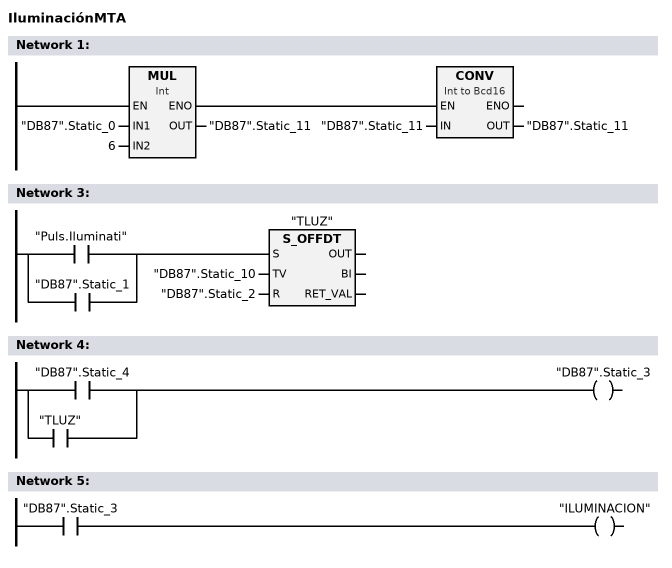
   RUNG wire#powerrail
      { S7_Templates := "SrcType := Int"; S7_GenerateENO := "TRUE" } Mul(in1 := "DB87".Static_0, in2 := 6, out => "DB87".Static_11)
      { S7_Templates := "[SrcType := Int, DestType := Bcd16]"; S7_GenerateENO := "TRUE" } Convert(in := "DB87".Static_11, out => "DB87".Static_11)
   END_RUNG
   // the same network as SCL:
   // ENO of a box is taken as its EN; it also drops when the box reports an error
   "DB87".Static_11 := "DB87".Static_0 * 6;
   "DB87".Static_11 := INT_TO_BCD16("DB87".Static_11);
END_REGION

REGION Network 2 (STL)
         L     12288;
         L     "DB87".Static_11;
         OW;
         T     "DB87".Static_10;
         NOP   0;
END_REGION

REGION Network 3
   RUNG wire#powerrail
      Contact( "Puls.Iluminati" )
      wire#w1
      S_OFFDT(T_NO := "TLUZ", TV := "DB87".Static_10, R := "DB87".Static_2, BI =>, RET_VAL =>)
   END_RUNG
   RUNG wire#powerrail
      Contact( "DB87".Static_1 )
   END_RUNG wire#w1
   // the same network as SCL:
   #_s5time1 := S_OFFDT(T_NO := "TLUZ",
                        S := "Puls.Iluminati" OR "DB87".Static_1,
                        TV := "DB87".Static_10,
                        R := "DB87".Static_2);
END_REGION

REGION Network 4
   RUNG wire#powerrail
      Contact( "DB87".Static_4 )
      wire#w1
      Coil( "DB87".Static_3 )
   END_RUNG
   RUNG wire#powerrail
      Contact( "TLUZ" )
   END_RUNG wire#w1
   // the same network as SCL:
   "DB87".Static_3 := "DB87".Static_4 OR "TLUZ";
END_REGION

REGION Network 5
   RUNG wire#powerrail
      Contact( "DB87".Static_3 )
      Coil( "ILUMINACION" )
   END_RUNG
   // the same network as SCL:
   "ILUMINACION" := "DB87".Static_3;
END_REGION
END_FUNCTION

// folder: OBs de fallas

ORGANIZATION_BLOCK "OB40"   // OB40, STL
{ S7_Optimized_Access := 'FALSE' }
VERSION : 0.0
BEGIN
END_ORGANIZATION_BLOCK

ORGANIZATION_BLOCK "Cycle Time Fault"   // OB80, STL
{ S7_Optimized_Access := 'FALSE' }
VERSION : 0.0
BEGIN
END_ORGANIZATION_BLOCK

ORGANIZATION_BLOCK "I/O Point Fault 1"   // OB82, LAD
{ S7_Optimized_Access := 'FALSE' }
VERSION : 0.1
BEGIN
END_ORGANIZATION_BLOCK

ORGANIZATION_BLOCK "OB83"   // OB83, STL
{ S7_Optimized_Access := 'FALSE' }
VERSION : 0.1
BEGIN
END_ORGANIZATION_BLOCK

ORGANIZATION_BLOCK "OB Not Loaded Fault"   // OB85, LAD
{ S7_Optimized_Access := 'FALSE' }
VERSION : 0.1
BEGIN
END_ORGANIZATION_BLOCK

ORGANIZATION_BLOCK "Fallo del bastidor"   // OB86, STL
{ S7_Optimized_Access := 'FALSE' }
VERSION : 0.1
BEGIN
END_ORGANIZATION_BLOCK

ORGANIZATION_BLOCK "Communication Fault"   // OB87, LAD
{ S7_Optimized_Access := 'FALSE' }
VERSION : 0.1
BEGIN
END_ORGANIZATION_BLOCK

ORGANIZATION_BLOCK "Complete Restart"   // OB100, LAD
{ S7_Optimized_Access := 'FALSE' }
VERSION : 0.1
BEGIN
END_ORGANIZATION_BLOCK

ORGANIZATION_BLOCK "Programming Error"   // OB121, LAD
{ S7_Optimized_Access := 'FALSE' }
VERSION : 0.1
BEGIN
END_ORGANIZATION_BLOCK

ORGANIZATION_BLOCK "Module Access Error"   // OB122, LAD
{ S7_Optimized_Access := 'FALSE' }
VERSION : 0.1
BEGIN
END_ORGANIZATION_BLOCK

// folder: Panel

FUNCTION_BLOCK "CHControlMotorPanelMTA"   // FB55, LAD
{ S7_Optimized_Access := 'FALSE' }
VERSION : 0.1
   VAR_TEMP   // added for the SCL form of the ladder/FBD networks
      _w1 : Bool;
   END_VAR
BEGIN

REGION Network 1
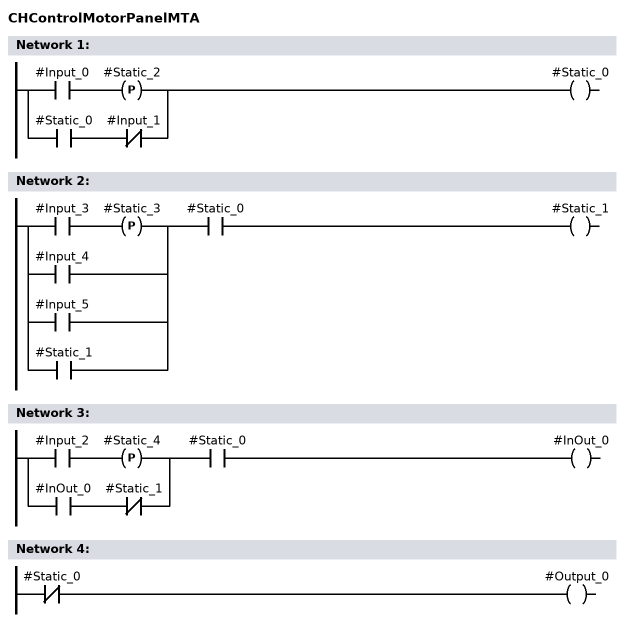
   RUNG wire#powerrail
      Contact( #Input_0 )
      P_Trig( #Static_2 )
      wire#w1
      Coil( #Static_0 )
   END_RUNG
   RUNG wire#powerrail
      Contact( #Static_0 )
      I_Contact( #Input_1 )
   END_RUNG wire#w1
   // the same network as SCL:
   #_w1 := #Input_0 AND NOT #Static_2;   // rising edge
   #Static_2 := #Input_0;
   #Static_0 := #_w1 OR (#Static_0 AND NOT #Input_1);
END_REGION

REGION Network 2
   RUNG wire#powerrail
      Contact( #Input_3 )
      P_Trig( #Static_3 )
      wire#w1
      Contact( #Static_0 )
      Coil( #Static_1 )
   END_RUNG
   RUNG wire#powerrail
      Contact( #Input_4 )
   END_RUNG wire#w1
   RUNG wire#powerrail
      Contact( #Input_5 )
   END_RUNG wire#w1
   RUNG wire#powerrail
      Contact( #Static_1 )
   END_RUNG wire#w1
   // the same network as SCL:
   #_w1 := #Input_3 AND NOT #Static_3;   // rising edge
   #Static_3 := #Input_3;
   #Static_1 := (#_w1 OR #Input_4 OR #Input_5 OR #Static_1) AND #Static_0;
END_REGION

REGION Network 3
   RUNG wire#powerrail
      Contact( #Input_2 )
      P_Trig( #Static_4 )
      wire#w1
      Contact( #Static_0 )
      Coil( #InOut_0 )
   END_RUNG
   RUNG wire#powerrail
      Contact( #InOut_0 )
      I_Contact( #Static_1 )
   END_RUNG wire#w1
   // the same network as SCL:
   #_w1 := #Input_2 AND NOT #Static_4;   // rising edge
   #Static_4 := #Input_2;
   #InOut_0 := (#_w1 OR (#InOut_0 AND NOT #Static_1)) AND #Static_0;
END_REGION

REGION Network 4
   RUNG wire#powerrail
      I_Contact( #Static_0 )
      Coil( #Output_0 )
   END_RUNG
   // the same network as SCL:
   #Output_0 := NOT #Static_0;
END_REGION
END_FUNCTION_BLOCK

FUNCTION "AnimaciónMTA" : Void   // FC2, LAD
{ S7_Optimized_Access := 'FALSE' }
VERSION : 0.1
   VAR_TEMP   // added for the SCL form of the ladder/FBD networks
      _w1 : Bool;
      _w2 : Bool;
   END_VAR
BEGIN

REGION Network 1
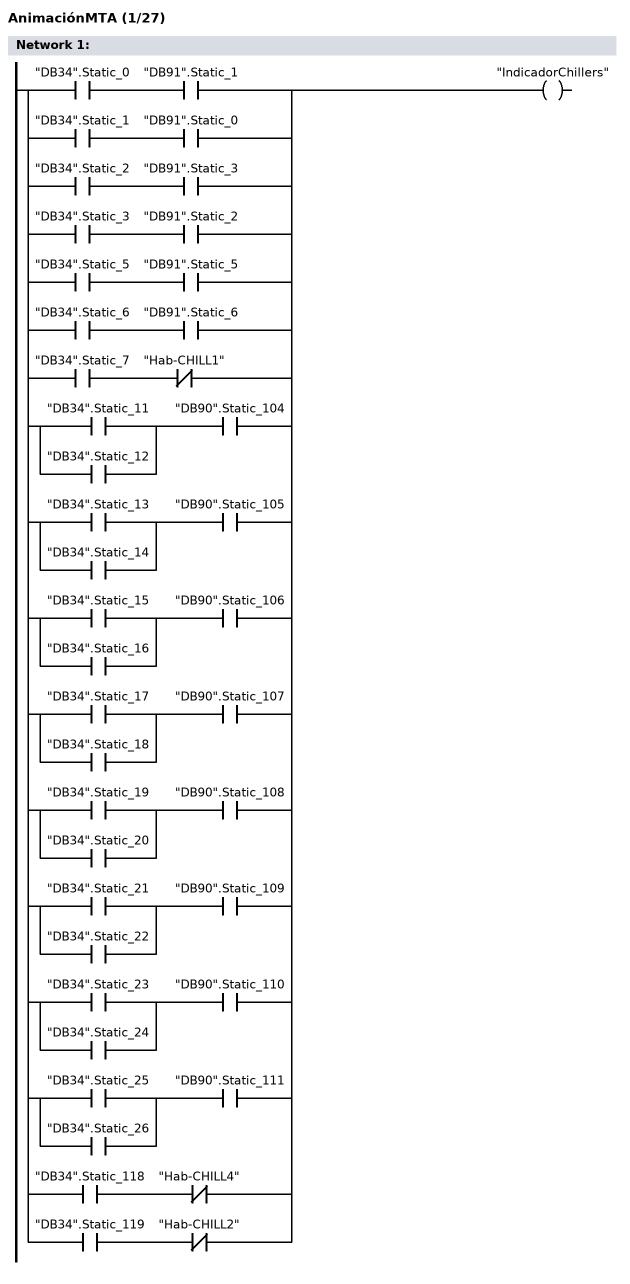
   RUNG wire#powerrail
      Contact( "DB34".Static_0 )
      Contact( "DB91".Static_1 )
      wire#w1
      Coil( "IndicadorChillers" )
   END_RUNG
   RUNG wire#powerrail
      Contact( "DB34".Static_1 )
      Contact( "DB91".Static_0 )
   END_RUNG wire#w1
   RUNG wire#powerrail
      Contact( "DB34".Static_2 )
      Contact( "DB91".Static_3 )
   END_RUNG wire#w1
   RUNG wire#powerrail
      Contact( "DB34".Static_3 )
      Contact( "DB91".Static_2 )
   END_RUNG wire#w1
   RUNG wire#powerrail
      Contact( "DB34".Static_5 )
      Contact( "DB91".Static_5 )
   END_RUNG wire#w1
   RUNG wire#powerrail
      Contact( "DB34".Static_6 )
      Contact( "DB91".Static_6 )
   END_RUNG wire#w1
   RUNG wire#powerrail
      Contact( "DB34".Static_7 )
      I_Contact( "Hab-CHILL1" )
   END_RUNG wire#w1
   RUNG wire#powerrail
      Contact( "DB34".Static_11 )
      wire#w2
      Contact( "DB90".Static_104 )
   END_RUNG wire#w1
   RUNG wire#powerrail
      Contact( "DB34".Static_12 )
   END_RUNG wire#w2
   RUNG wire#powerrail
      Contact( "DB34".Static_13 )
      wire#w3
      Contact( "DB90".Static_105 )
   END_RUNG wire#w1
   RUNG wire#powerrail
      Contact( "DB34".Static_14 )
   END_RUNG wire#w3
   RUNG wire#powerrail
      Contact( "DB34".Static_15 )
      wire#w4
      Contact( "DB90".Static_106 )
   END_RUNG wire#w1
   RUNG wire#powerrail
      Contact( "DB34".Static_16 )
   END_RUNG wire#w4
   RUNG wire#powerrail
      Contact( "DB34".Static_17 )
      wire#w5
      Contact( "DB90".Static_107 )
   END_RUNG wire#w1
   RUNG wire#powerrail
      Contact( "DB34".Static_18 )
   END_RUNG wire#w5
   RUNG wire#powerrail
      Contact( "DB34".Static_19 )
      wire#w6
      Contact( "DB90".Static_108 )
   END_RUNG wire#w1
   RUNG wire#powerrail
      Contact( "DB34".Static_20 )
   END_RUNG wire#w6
   RUNG wire#powerrail
      Contact( "DB34".Static_21 )
      wire#w7
      Contact( "DB90".Static_109 )
   END_RUNG wire#w1
   RUNG wire#powerrail
      Contact( "DB34".Static_22 )
   END_RUNG wire#w7
   RUNG wire#powerrail
      Contact( "DB34".Static_23 )
      wire#w8
      Contact( "DB90".Static_110 )
   END_RUNG wire#w1
   RUNG wire#powerrail
      Contact( "DB34".Static_24 )
   END_RUNG wire#w8
   RUNG wire#powerrail
      Contact( "DB34".Static_25 )
      wire#w9
      Contact( "DB90".Static_111 )
   END_RUNG wire#w1
   RUNG wire#powerrail
      Contact( "DB34".Static_26 )
   END_RUNG wire#w9
   RUNG wire#powerrail
      Contact( "DB34".Static_118 )
      I_Contact( "Hab-CHILL4" )
   END_RUNG wire#w1
   RUNG wire#powerrail
      Contact( "DB34".Static_119 )
      I_Contact( "Hab-CHILL2" )
   END_RUNG wire#w1
   // the same network as SCL:
   "IndicadorChillers" := ("DB34".Static_0 AND "DB91".Static_1) OR ("DB34".Static_1 AND "DB91".Static_0) OR ("DB34".Static_2 AND "DB91".Static_3) OR ("DB34".Static_3 AND "DB91".Static_2) OR ("DB34".Static_5 AND "DB91".Static_5) OR ("DB34".Static_6 AND "DB91".Static_6) OR ("DB34".Static_7 AND NOT "Hab-CHILL1") OR (("DB34".Static_11 OR "DB34".Static_12) AND "DB90".Static_104) OR (("DB34".Static_13 OR "DB34".Static_14) AND "DB90".Static_105) OR (("DB34".Static_15 OR "DB34".Static_16) AND "DB90".Static_106) OR (("DB34".Static_17 OR "DB34".Static_18) AND "DB90".Static_107) OR (("DB34".Static_19 OR "DB34".Static_20) AND "DB90".Static_108) OR (("DB34".Static_21 OR "DB34".Static_22) AND "DB90".Static_109) OR (("DB34".Static_23 OR "DB34".Static_24) AND "DB90".Static_110) OR (("DB34".Static_25 OR "DB34".Static_26) AND "DB90".Static_111) OR ("DB34".Static_118 AND NOT "Hab-CHILL4") OR ("DB34".Static_119 AND NOT "Hab-CHILL2");
END_REGION

REGION Network 2
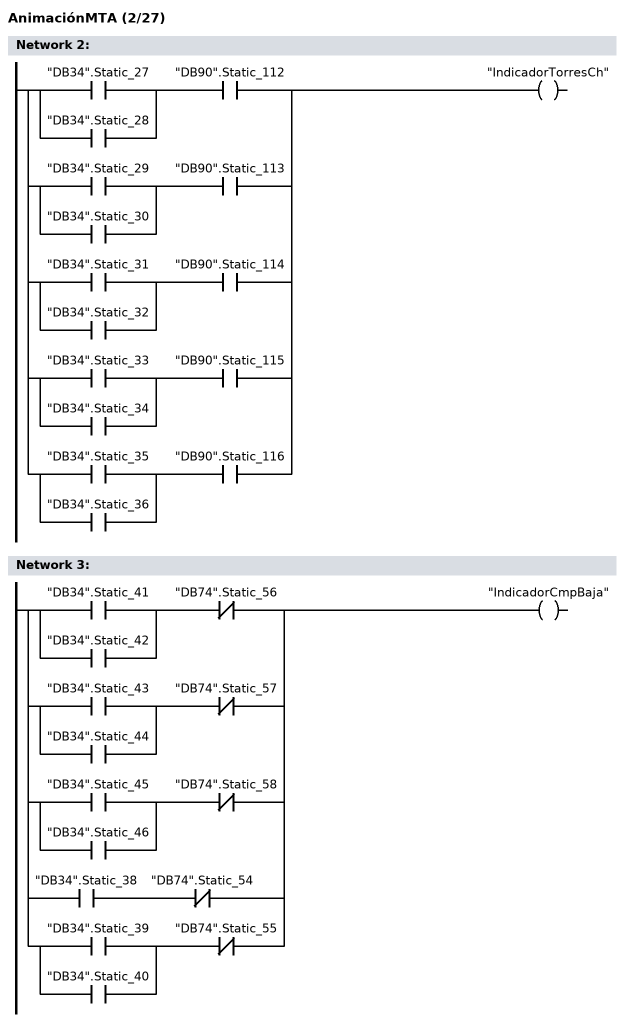
   RUNG wire#powerrail
      Contact( "DB34".Static_27 )
      wire#w1
      Contact( "DB90".Static_112 )
      wire#w2
      Coil( "IndicadorTorresCh" )
   END_RUNG
   RUNG wire#powerrail
      Contact( "DB34".Static_28 )
   END_RUNG wire#w1
   RUNG wire#powerrail
      Contact( "DB34".Static_29 )
      wire#w3
      Contact( "DB90".Static_113 )
   END_RUNG wire#w2
   RUNG wire#powerrail
      Contact( "DB34".Static_30 )
   END_RUNG wire#w3
   RUNG wire#powerrail
      Contact( "DB34".Static_31 )
      wire#w4
      Contact( "DB90".Static_114 )
   END_RUNG wire#w2
   RUNG wire#powerrail
      Contact( "DB34".Static_32 )
   END_RUNG wire#w4
   RUNG wire#powerrail
      Contact( "DB34".Static_33 )
      wire#w5
      Contact( "DB90".Static_115 )
   END_RUNG wire#w2
   RUNG wire#powerrail
      Contact( "DB34".Static_34 )
   END_RUNG wire#w5
   RUNG wire#powerrail
      Contact( "DB34".Static_35 )
      wire#w6
      Contact( "DB90".Static_116 )
   END_RUNG wire#w2
   RUNG wire#powerrail
      Contact( "DB34".Static_36 )
   END_RUNG wire#w6
   // the same network as SCL:
   "IndicadorTorresCh" := (("DB34".Static_27 OR "DB34".Static_28) AND "DB90".Static_112) OR (("DB34".Static_29 OR "DB34".Static_30) AND "DB90".Static_113) OR (("DB34".Static_31 OR "DB34".Static_32) AND "DB90".Static_114) OR (("DB34".Static_33 OR "DB34".Static_34) AND "DB90".Static_115) OR (("DB34".Static_35 OR "DB34".Static_36) AND "DB90".Static_116);
END_REGION

REGION Network 3
   RUNG wire#powerrail
      Contact( "DB34".Static_41 )
      wire#w1
      I_Contact( "DB74".Static_56 )
      wire#w2
      Coil( "IndicadorCmpBaja" )
   END_RUNG
   RUNG wire#powerrail
      Contact( "DB34".Static_42 )
   END_RUNG wire#w1
   RUNG wire#powerrail
      Contact( "DB34".Static_43 )
      wire#w3
      I_Contact( "DB74".Static_57 )
   END_RUNG wire#w2
   RUNG wire#powerrail
      Contact( "DB34".Static_44 )
   END_RUNG wire#w3
   RUNG wire#powerrail
      Contact( "DB34".Static_45 )
      wire#w4
      I_Contact( "DB74".Static_58 )
   END_RUNG wire#w2
   RUNG wire#powerrail
      Contact( "DB34".Static_46 )
   END_RUNG wire#w4
   RUNG wire#powerrail
      Contact( "DB34".Static_38 )
      I_Contact( "DB74".Static_54 )
   END_RUNG wire#w2
   RUNG wire#powerrail
      Contact( "DB34".Static_39 )
      wire#w5
      I_Contact( "DB74".Static_55 )
   END_RUNG wire#w2
   RUNG wire#powerrail
      Contact( "DB34".Static_40 )
   END_RUNG wire#w5
   // the same network as SCL:
   "IndicadorCmpBaja" := (("DB34".Static_41 OR "DB34".Static_42) AND NOT "DB74".Static_56) OR (("DB34".Static_43 OR "DB34".Static_44) AND NOT "DB74".Static_57) OR (("DB34".Static_45 OR "DB34".Static_46) AND NOT "DB74".Static_58) OR ("DB34".Static_38 AND NOT "DB74".Static_54) OR (("DB34".Static_39 OR "DB34".Static_40) AND NOT "DB74".Static_55);
END_REGION

REGION Network 4
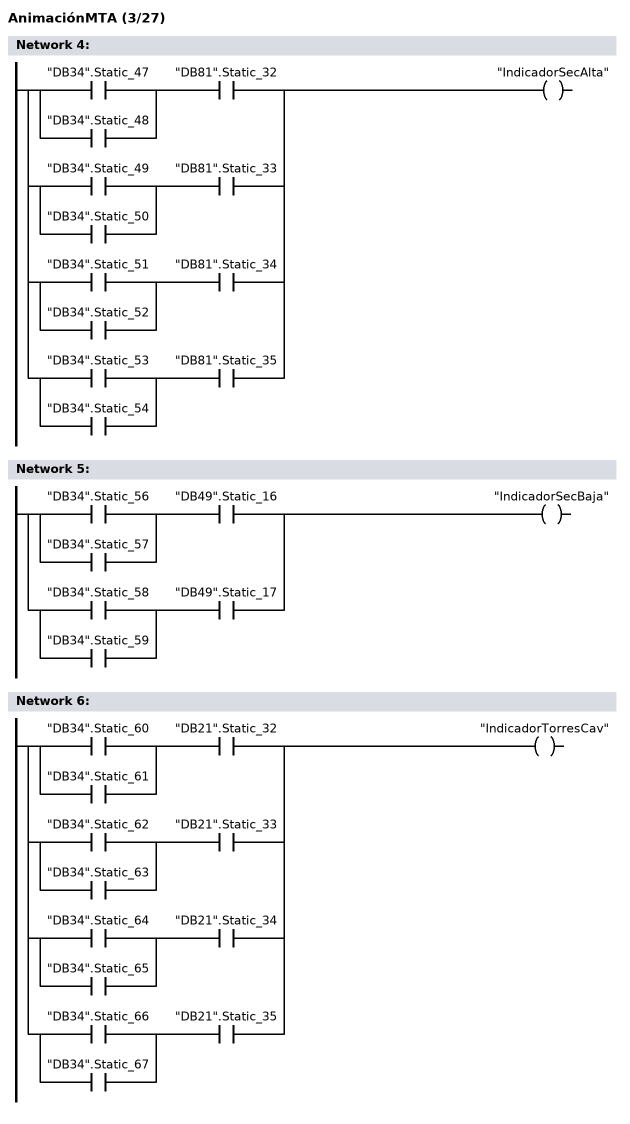
   RUNG wire#powerrail
      Contact( "DB34".Static_47 )
      wire#w1
      Contact( "DB81".Static_32 )
      wire#w2
      Coil( "IndicadorSecAlta" )
   END_RUNG
   RUNG wire#powerrail
      Contact( "DB34".Static_48 )
   END_RUNG wire#w1
   RUNG wire#powerrail
      Contact( "DB34".Static_49 )
      wire#w3
      Contact( "DB81".Static_33 )
   END_RUNG wire#w2
   RUNG wire#powerrail
      Contact( "DB34".Static_50 )
   END_RUNG wire#w3
   RUNG wire#powerrail
      Contact( "DB34".Static_51 )
      wire#w4
      Contact( "DB81".Static_34 )
   END_RUNG wire#w2
   RUNG wire#powerrail
      Contact( "DB34".Static_52 )
   END_RUNG wire#w4
   RUNG wire#powerrail
      Contact( "DB34".Static_53 )
      wire#w5
      Contact( "DB81".Static_35 )
   END_RUNG wire#w2
   RUNG wire#powerrail
      Contact( "DB34".Static_54 )
   END_RUNG wire#w5
   // the same network as SCL:
   "IndicadorSecAlta" := (("DB34".Static_47 OR "DB34".Static_48) AND "DB81".Static_32) OR (("DB34".Static_49 OR "DB34".Static_50) AND "DB81".Static_33) OR (("DB34".Static_51 OR "DB34".Static_52) AND "DB81".Static_34) OR (("DB34".Static_53 OR "DB34".Static_54) AND "DB81".Static_35);
END_REGION

REGION Network 5
   RUNG wire#powerrail
      Contact( "DB34".Static_56 )
      wire#w1
      Contact( "DB49".Static_16 )
      wire#w2
      Coil( "IndicadorSecBaja" )
   END_RUNG
   RUNG wire#powerrail
      Contact( "DB34".Static_57 )
   END_RUNG wire#w1
   RUNG wire#powerrail
      Contact( "DB34".Static_58 )
      wire#w3
      Contact( "DB49".Static_17 )
   END_RUNG wire#w2
   RUNG wire#powerrail
      Contact( "DB34".Static_59 )
   END_RUNG wire#w3
   // the same network as SCL:
   "IndicadorSecBaja" := (("DB34".Static_56 OR "DB34".Static_57) AND "DB49".Static_16) OR (("DB34".Static_58 OR "DB34".Static_59) AND "DB49".Static_17);
END_REGION

REGION Network 6
   RUNG wire#powerrail
      Contact( "DB34".Static_60 )
      wire#w1
      Contact( "DB21".Static_32 )
      wire#w2
      Coil( "IndicadorTorresCav" )
   END_RUNG
   RUNG wire#powerrail
      Contact( "DB34".Static_61 )
   END_RUNG wire#w1
   RUNG wire#powerrail
      Contact( "DB34".Static_62 )
      wire#w3
      Contact( "DB21".Static_33 )
   END_RUNG wire#w2
   RUNG wire#powerrail
      Contact( "DB34".Static_63 )
   END_RUNG wire#w3
   RUNG wire#powerrail
      Contact( "DB34".Static_64 )
      wire#w4
      Contact( "DB21".Static_34 )
   END_RUNG wire#w2
   RUNG wire#powerrail
      Contact( "DB34".Static_65 )
   END_RUNG wire#w4
   RUNG wire#powerrail
      Contact( "DB34".Static_66 )
      wire#w5
      Contact( "DB21".Static_35 )
   END_RUNG wire#w2
   RUNG wire#powerrail
      Contact( "DB34".Static_67 )
   END_RUNG wire#w5
   // the same network as SCL:
   "IndicadorTorresCav" := (("DB34".Static_60 OR "DB34".Static_61) AND "DB21".Static_32) OR (("DB34".Static_62 OR "DB34".Static_63) AND "DB21".Static_33) OR (("DB34".Static_64 OR "DB34".Static_65) AND "DB21".Static_34) OR (("DB34".Static_66 OR "DB34".Static_67) AND "DB21".Static_35);
END_REGION

REGION Network 7
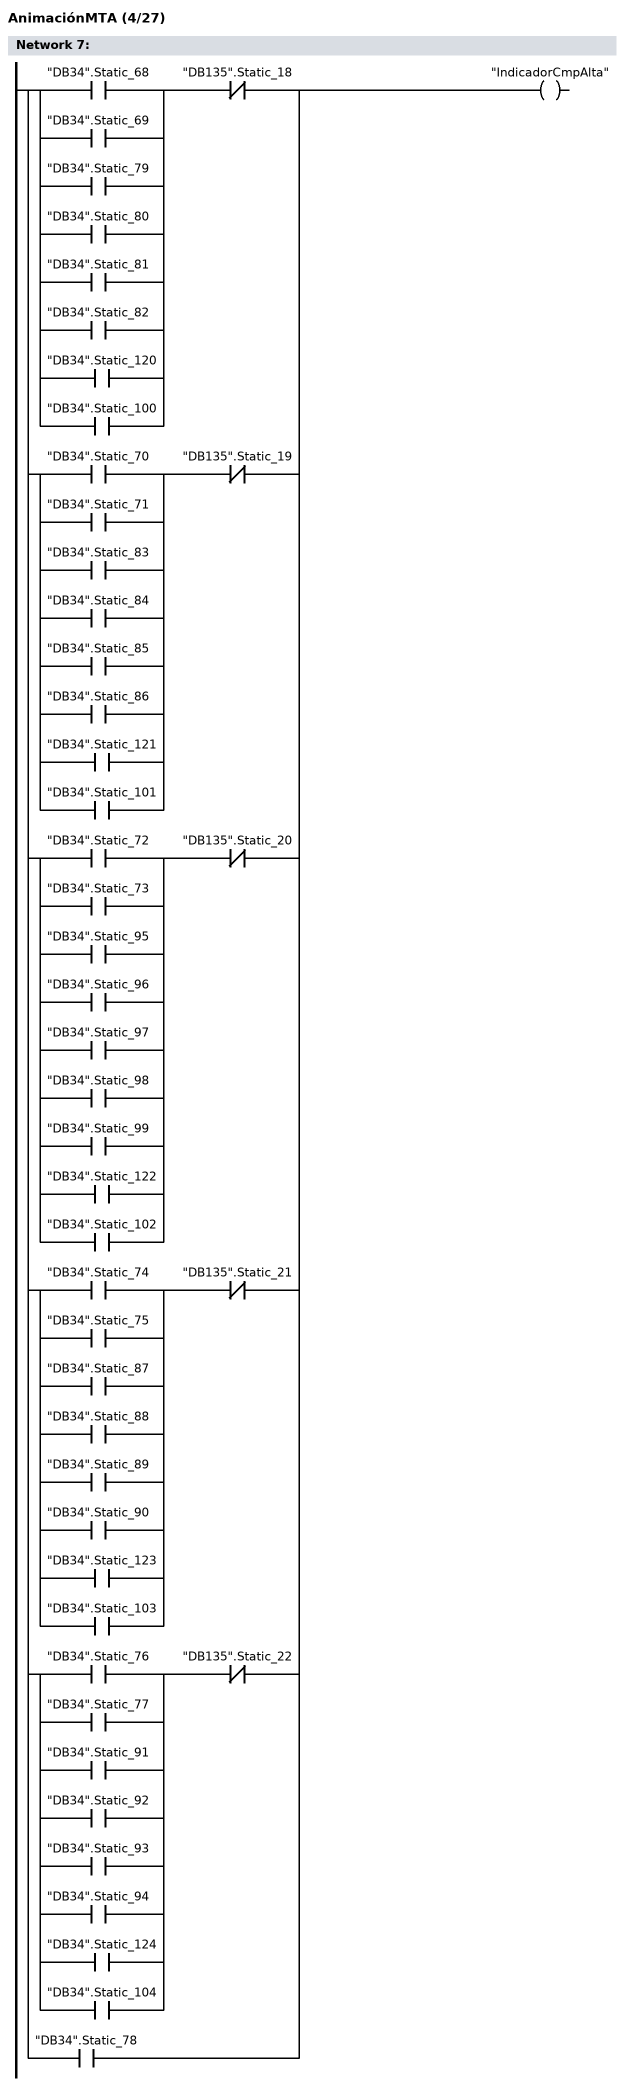
   RUNG wire#powerrail
      Contact( "DB34".Static_68 )
      wire#w1
      I_Contact( "DB135".Static_18 )
      wire#w2
      Coil( "IndicadorCmpAlta" )
   END_RUNG
   RUNG wire#powerrail
      Contact( "DB34".Static_69 )
   END_RUNG wire#w1
   RUNG wire#powerrail
      Contact( "DB34".Static_79 )
   END_RUNG wire#w1
   RUNG wire#powerrail
      Contact( "DB34".Static_80 )
   END_RUNG wire#w1
   RUNG wire#powerrail
      Contact( "DB34".Static_81 )
   END_RUNG wire#w1
   RUNG wire#powerrail
      Contact( "DB34".Static_82 )
   END_RUNG wire#w1
   RUNG wire#powerrail
      Contact( "DB34".Static_120 )
   END_RUNG wire#w1
   RUNG wire#powerrail
      Contact( "DB34".Static_100 )
   END_RUNG wire#w1
   RUNG wire#powerrail
      Contact( "DB34".Static_70 )
      wire#w3
      I_Contact( "DB135".Static_19 )
   END_RUNG wire#w2
   RUNG wire#powerrail
      Contact( "DB34".Static_71 )
   END_RUNG wire#w3
   RUNG wire#powerrail
      Contact( "DB34".Static_83 )
   END_RUNG wire#w3
   RUNG wire#powerrail
      Contact( "DB34".Static_84 )
   END_RUNG wire#w3
   RUNG wire#powerrail
      Contact( "DB34".Static_85 )
   END_RUNG wire#w3
   RUNG wire#powerrail
      Contact( "DB34".Static_86 )
   END_RUNG wire#w3
   RUNG wire#powerrail
      Contact( "DB34".Static_121 )
   END_RUNG wire#w3
   RUNG wire#powerrail
      Contact( "DB34".Static_101 )
   END_RUNG wire#w3
   RUNG wire#powerrail
      Contact( "DB34".Static_72 )
      wire#w4
      I_Contact( "DB135".Static_20 )
   END_RUNG wire#w2
   RUNG wire#powerrail
      Contact( "DB34".Static_73 )
   END_RUNG wire#w4
   RUNG wire#powerrail
      Contact( "DB34".Static_95 )
   END_RUNG wire#w4
   RUNG wire#powerrail
      Contact( "DB34".Static_96 )
   END_RUNG wire#w4
   RUNG wire#powerrail
      Contact( "DB34".Static_97 )
   END_RUNG wire#w4
   RUNG wire#powerrail
      Contact( "DB34".Static_98 )
   END_RUNG wire#w4
   RUNG wire#powerrail
      Contact( "DB34".Static_99 )
   END_RUNG wire#w4
   RUNG wire#powerrail
      Contact( "DB34".Static_122 )
   END_RUNG wire#w4
   RUNG wire#powerrail
      Contact( "DB34".Static_102 )
   END_RUNG wire#w4
   RUNG wire#powerrail
      Contact( "DB34".Static_74 )
      wire#w5
      I_Contact( "DB135".Static_21 )
   END_RUNG wire#w2
   RUNG wire#powerrail
      Contact( "DB34".Static_75 )
   END_RUNG wire#w5
   RUNG wire#powerrail
      Contact( "DB34".Static_87 )
   END_RUNG wire#w5
   RUNG wire#powerrail
      Contact( "DB34".Static_88 )
   END_RUNG wire#w5
   RUNG wire#powerrail
      Contact( "DB34".Static_89 )
   END_RUNG wire#w5
   RUNG wire#powerrail
      Contact( "DB34".Static_90 )
   END_RUNG wire#w5
   RUNG wire#powerrail
      Contact( "DB34".Static_123 )
   END_RUNG wire#w5
   RUNG wire#powerrail
      Contact( "DB34".Static_103 )
   END_RUNG wire#w5
   RUNG wire#powerrail
      Contact( "DB34".Static_76 )
      wire#w6
      I_Contact( "DB135".Static_22 )
   END_RUNG wire#w2
   RUNG wire#powerrail
      Contact( "DB34".Static_77 )
   END_RUNG wire#w6
   RUNG wire#powerrail
      Contact( "DB34".Static_91 )
   END_RUNG wire#w6
   RUNG wire#powerrail
      Contact( "DB34".Static_92 )
   END_RUNG wire#w6
   RUNG wire#powerrail
      Contact( "DB34".Static_93 )
   END_RUNG wire#w6
   RUNG wire#powerrail
      Contact( "DB34".Static_94 )
   END_RUNG wire#w6
   RUNG wire#powerrail
      Contact( "DB34".Static_124 )
   END_RUNG wire#w6
   RUNG wire#powerrail
      Contact( "DB34".Static_104 )
   END_RUNG wire#w6
   RUNG wire#powerrail
      Contact( "DB34".Static_78 )
   END_RUNG wire#w2
   // the same network as SCL:
   "IndicadorCmpAlta" := (("DB34".Static_68 OR "DB34".Static_69 OR "DB34".Static_79 OR "DB34".Static_80 OR "DB34".Static_81 OR "DB34".Static_82 OR "DB34".Static_120 OR "DB34".Static_100) AND NOT "DB135".Static_18) OR (("DB34".Static_70 OR "DB34".Static_71 OR "DB34".Static_83 OR "DB34".Static_84 OR "DB34".Static_85 OR "DB34".Static_86 OR "DB34".Static_121 OR "DB34".Static_101) AND NOT "DB135".Static_19) OR (("DB34".Static_72 OR "DB34".Static_73 OR "DB34".Static_95 OR "DB34".Static_96 OR "DB34".Static_97 OR "DB34".Static_98 OR "DB34".Static_99 OR "DB34".Static_122 OR "DB34".Static_102) AND NOT "DB135".Static_20) OR (("DB34".Static_74 OR "DB34".Static_75 OR "DB34".Static_87 OR "DB34".Static_88 OR "DB34".Static_89 OR "DB34".Static_90 OR "DB34".Static_123 OR "DB34".Static_103) AND NOT "DB135".Static_21) OR (("DB34".Static_76 OR "DB34".Static_77 OR "DB34".Static_91 OR "DB34".Static_92 OR "DB34".Static_93 OR "DB34".Static_94 OR "DB34".Static_124 OR "DB34".Static_104) AND NOT "DB135".Static_22) OR "DB34".Static_78;
END_REGION

REGION Network 8
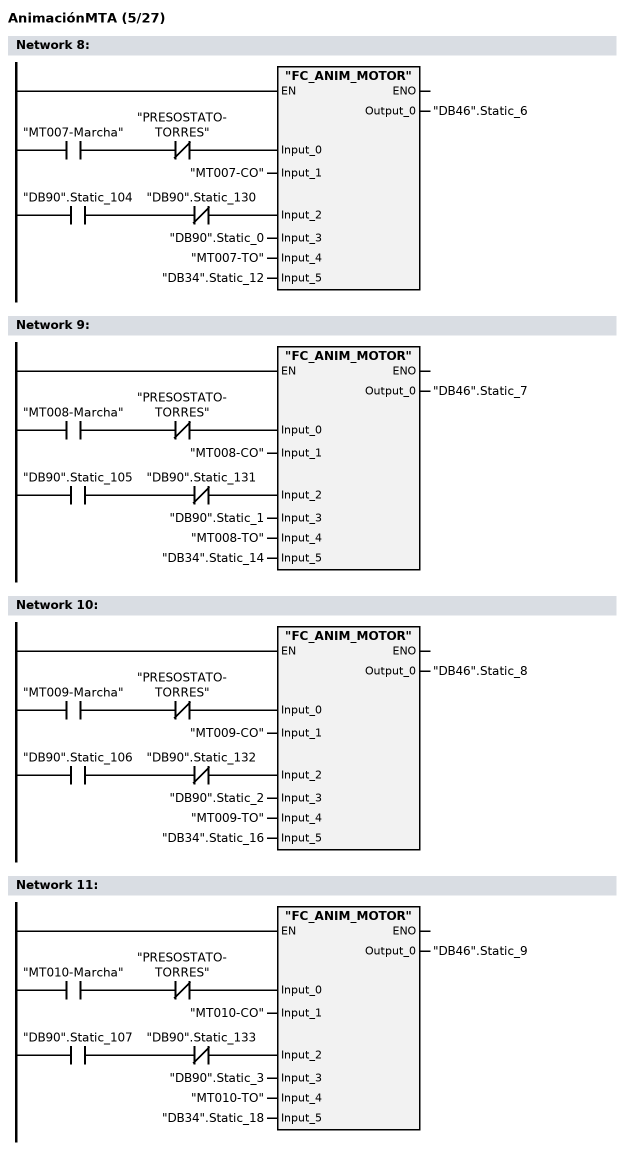
   RUNG wire#powerrail
      "FC_ANIM_MOTOR"(Input_1 := "MT007-CO", Input_3 := "DB90".Static_0, Input_4 := "MT007-TO", Input_5 := "DB34".Static_12, Output_0 => "DB46".Static_6, Input_0 := wire#w1, Input_2 := wire#w2)
   END_RUNG
   RUNG wire#powerrail
      Contact( "MT007-Marcha" )
      I_Contact( "PRESOSTATO-TORRES" )
   END_RUNG wire#w1
   RUNG wire#powerrail
      Contact( "DB90".Static_104 )
      I_Contact( "DB90".Static_130 )
   END_RUNG wire#w2
   // the same network as SCL:
   "FC_ANIM_MOTOR"(Input_0 := "MT007-Marcha" AND NOT "PRESOSTATO-TORRES",
                   Input_1 := "MT007-CO",
                   Input_2 := "DB90".Static_104 AND NOT "DB90".Static_130,
                   Input_3 := "DB90".Static_0,
                   Input_4 := "MT007-TO",
                   Input_5 := "DB34".Static_12,
                   Output_0 => "DB46".Static_6);
END_REGION

REGION Network 9
   RUNG wire#powerrail
      "FC_ANIM_MOTOR"(Input_1 := "MT008-CO", Input_3 := "DB90".Static_1, Input_4 := "MT008-TO", Input_5 := "DB34".Static_14, Output_0 => "DB46".Static_7, Input_0 := wire#w1, Input_2 := wire#w2)
   END_RUNG
   RUNG wire#powerrail
      Contact( "MT008-Marcha" )
      I_Contact( "PRESOSTATO-TORRES" )
   END_RUNG wire#w1
   RUNG wire#powerrail
      Contact( "DB90".Static_105 )
      I_Contact( "DB90".Static_131 )
   END_RUNG wire#w2
   // the same network as SCL:
   "FC_ANIM_MOTOR"(Input_0 := "MT008-Marcha" AND NOT "PRESOSTATO-TORRES",
                   Input_1 := "MT008-CO",
                   Input_2 := "DB90".Static_105 AND NOT "DB90".Static_131,
                   Input_3 := "DB90".Static_1,
                   Input_4 := "MT008-TO",
                   Input_5 := "DB34".Static_14,
                   Output_0 => "DB46".Static_7);
END_REGION

REGION Network 10
   RUNG wire#powerrail
      "FC_ANIM_MOTOR"(Input_1 := "MT009-CO", Input_3 := "DB90".Static_2, Input_4 := "MT009-TO", Input_5 := "DB34".Static_16, Output_0 => "DB46".Static_8, Input_0 := wire#w1, Input_2 := wire#w2)
   END_RUNG
   RUNG wire#powerrail
      Contact( "MT009-Marcha" )
      I_Contact( "PRESOSTATO-TORRES" )
   END_RUNG wire#w1
   RUNG wire#powerrail
      Contact( "DB90".Static_106 )
      I_Contact( "DB90".Static_132 )
   END_RUNG wire#w2
   // the same network as SCL:
   "FC_ANIM_MOTOR"(Input_0 := "MT009-Marcha" AND NOT "PRESOSTATO-TORRES",
                   Input_1 := "MT009-CO",
                   Input_2 := "DB90".Static_106 AND NOT "DB90".Static_132,
                   Input_3 := "DB90".Static_2,
                   Input_4 := "MT009-TO",
                   Input_5 := "DB34".Static_16,
                   Output_0 => "DB46".Static_8);
END_REGION

REGION Network 11
   RUNG wire#powerrail
      "FC_ANIM_MOTOR"(Input_1 := "MT010-CO", Input_3 := "DB90".Static_3, Input_4 := "MT010-TO", Input_5 := "DB34".Static_18, Output_0 => "DB46".Static_9, Input_0 := wire#w1, Input_2 := wire#w2)
   END_RUNG
   RUNG wire#powerrail
      Contact( "MT010-Marcha" )
      I_Contact( "PRESOSTATO-TORRES" )
   END_RUNG wire#w1
   RUNG wire#powerrail
      Contact( "DB90".Static_107 )
      I_Contact( "DB90".Static_133 )
   END_RUNG wire#w2
   // the same network as SCL:
   "FC_ANIM_MOTOR"(Input_0 := "MT010-Marcha" AND NOT "PRESOSTATO-TORRES",
                   Input_1 := "MT010-CO",
                   Input_2 := "DB90".Static_107 AND NOT "DB90".Static_133,
                   Input_3 := "DB90".Static_3,
                   Input_4 := "MT010-TO",
                   Input_5 := "DB34".Static_18,
                   Output_0 => "DB46".Static_9);
END_REGION

REGION Network 12
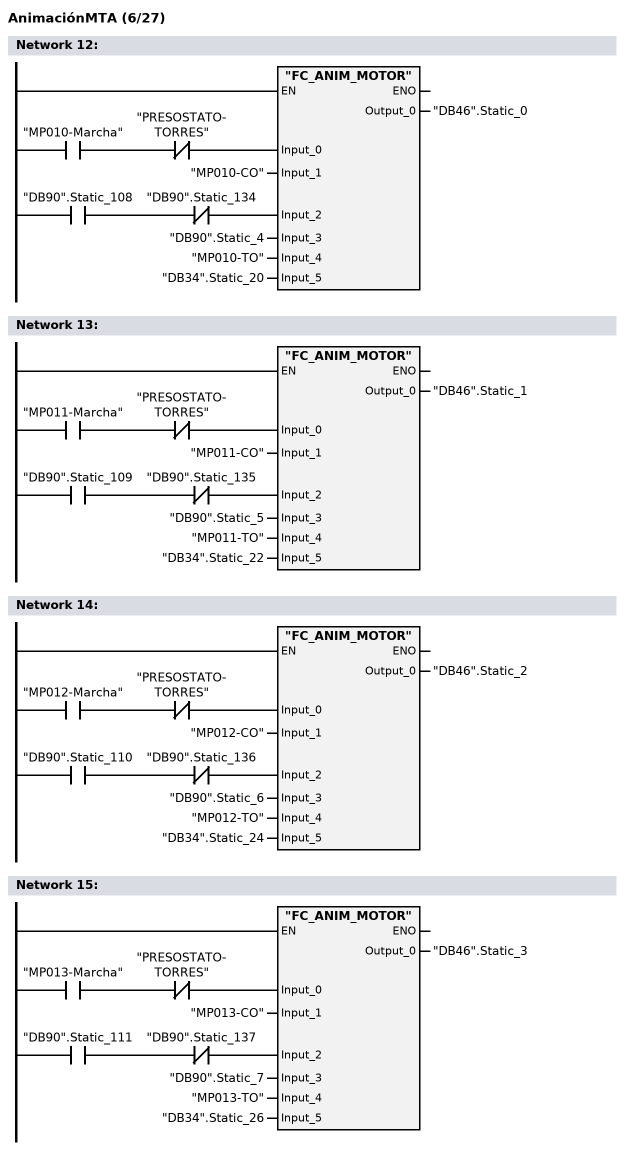
   RUNG wire#powerrail
      "FC_ANIM_MOTOR"(Input_1 := "MP010-CO", Input_3 := "DB90".Static_4, Input_4 := "MP010-TO", Input_5 := "DB34".Static_20, Output_0 => "DB46".Static_0, Input_0 := wire#w1, Input_2 := wire#w2)
   END_RUNG
   RUNG wire#powerrail
      Contact( "MP010-Marcha" )
      I_Contact( "PRESOSTATO-TORRES" )
   END_RUNG wire#w1
   RUNG wire#powerrail
      Contact( "DB90".Static_108 )
      I_Contact( "DB90".Static_134 )
   END_RUNG wire#w2
   // the same network as SCL:
   "FC_ANIM_MOTOR"(Input_0 := "MP010-Marcha" AND NOT "PRESOSTATO-TORRES",
                   Input_1 := "MP010-CO",
                   Input_2 := "DB90".Static_108 AND NOT "DB90".Static_134,
                   Input_3 := "DB90".Static_4,
                   Input_4 := "MP010-TO",
                   Input_5 := "DB34".Static_20,
                   Output_0 => "DB46".Static_0);
END_REGION

REGION Network 13
   RUNG wire#powerrail
      "FC_ANIM_MOTOR"(Input_1 := "MP011-CO", Input_3 := "DB90".Static_5, Input_4 := "MP011-TO", Input_5 := "DB34".Static_22, Output_0 => "DB46".Static_1, Input_0 := wire#w1, Input_2 := wire#w2)
   END_RUNG
   RUNG wire#powerrail
      Contact( "MP011-Marcha" )
      I_Contact( "PRESOSTATO-TORRES" )
   END_RUNG wire#w1
   RUNG wire#powerrail
      Contact( "DB90".Static_109 )
      I_Contact( "DB90".Static_135 )
   END_RUNG wire#w2
   // the same network as SCL:
   "FC_ANIM_MOTOR"(Input_0 := "MP011-Marcha" AND NOT "PRESOSTATO-TORRES",
                   Input_1 := "MP011-CO",
                   Input_2 := "DB90".Static_109 AND NOT "DB90".Static_135,
                   Input_3 := "DB90".Static_5,
                   Input_4 := "MP011-TO",
                   Input_5 := "DB34".Static_22,
                   Output_0 => "DB46".Static_1);
END_REGION
